HMI tags "xAI"
   "AIx_DB_Level_Use_RTD" : Bool = PLC AIx_DB.Level.Use.RTD AT %DB202.DBX156.0, 1 s
   "AIx_DB_Level_Use_Filter" : Bool = PLC AIx_DB.Level.Use.Filter AT %DB202.DBX156.1, 1 s
   "AIx_DB_Level_Timers_SC_SP" : Int = PLC AIx_DB.Level.Timers.SC.SP AT %DB202.DBW246, 1 s
   "AIx_DB_Level_Timers_NC_SP" : Int = PLC AIx_DB.Level.Timers.NC.SP AT %DB202.DBW240, 1 s
   "AIx_DB_Level_Timers_LL_SP" : Int = PLC AIx_DB.Level.Timers.LL.SP AT %DB202.DBW270, 1 s
   "AIx_DB_Level_Timers_L_SP" : Int = PLC AIx_DB.Level.Timers.L.SP AT %DB202.DBW264, 1 s
   "AIx_DB_Level_Timers_HH_SP" : Int = PLC AIx_DB.Level.Timers.HH.SP AT %DB202.DBW252, 1 s
   "AIx_DB_Level_Timers_H_SP" : Int = PLC AIx_DB.Level.Timers.H.SP AT %DB202.DBW258, 1 s
   "AIx_DB_Level_SP_SC" : Real = PLC AIx_DB.Level.SP.SC AT %DB202.DBD220, 1 s
   "AIx_DB_Level_SP_NC" : Real = PLC AIx_DB.Level.SP.NC AT %DB202.DBD216, 1 s
   "AIx_DB_Level_SP_LL" : Real = PLC AIx_DB.Level.SP.LL AT %DB202.DBD236, 1 s
   "AIx_DB_Level_SP_L" : Real = PLC AIx_DB.Level.SP.L AT %DB202.DBD232, 1 s
   "AIx_DB_Level_SP_HH" : Real = PLC AIx_DB.Level.SP.HH AT %DB202.DBD224, 1 s
   "AIx_DB_Level_SP_H" : Real = PLC AIx_DB.Level.SP.H AT %DB202.DBD228, 1 s
   "AIx_DB_Level_Signal" : Int = PLC AIx_DB.Level.Signal AT %DB202.DBW140, 1 s
   "AIx_DB_Level_RTD_c" : Real = PLC AIx_DB.Level.RTD_c AT %DB202.DBD170, 1 s
   "AIx_DB_Level_Result" : Real = PLC AIx_DB.Level.Result AT %DB202.DBD146, 1 s
   "AIx_DB_Level_Filter_SP" : Real = PLC AIx_DB.Level.Filter.SP AT %DB202.DBD178, 1 s
   "AIx_DB_Level_Converter_Min_Out" : Real = PLC AIx_DB.Level.Converter.Min_Out AT %DB202.DBD208, 1 s
   "AIx_DB_Level_Converter_Min_In" : Real = PLC AIx_DB.Level.Converter.Min_In AT %DB202.DBD200, 1 s
   "AIx_DB_Level_Converter_Max_Out" : Real = PLC AIx_DB.Level.Converter.Max_Out AT %DB202.DBD212, 1 s
   "AIx_DB_Level_Converter_Max_In" : Real = PLC AIx_DB.Level.Converter.Max_In AT %DB202.DBD204, 1 s
   "AIx_DB_Level_CMD_Start_M" : Bool = PLC AIx_DB.Level.CMD.Start_M AT %DB202.DBX150.2, 1 s
   "AIx_DB_Level_CMD_Start_A" : Bool = PLC AIx_DB.Level.CMD.Start_A AT %DB202.DBX150.1, 1 s
   "AIx_DB_Level_CMD_Hand" : Bool = PLC AIx_DB.Level.CMD.Hand AT %DB202.DBX150.0, 1 s
   "AIx_DB_Level_CMD_Alarm" : Bool = PLC AIx_DB.Level.CMD.Alarm AT %DB202.DBX151.0, 1 s
   "AIx_DB_Level_Calibration" : Real = PLC AIx_DB.Level.Calibration AT %DB202.DBD174, 1 s
   "AIx_DB_Level_Alarm" : Word = PLC AIx_DB.Level.Alarm AT %DB202.DBW278, 1 s
   "AIx_DB_FlowMeter_Use_RTD" : Bool = PLC AIx_DB.FlowMeter.Use.RTD AT %DB202.DBX16.0, 1 s
   "AIx_DB_FlowMeter_Use_Filter" : Bool = PLC AIx_DB.FlowMeter.Use.Filter AT %DB202.DBX16.1, 1 s
   "AIx_DB_FlowMeter_Timers_SC_SP" : Int = PLC AIx_DB.FlowMeter.Timers.SC.SP AT %DB202.DBW106, 1 s
   "AIx_DB_FlowMeter_Timers_NC_SP" : Int = PLC AIx_DB.FlowMeter.Timers.NC.SP AT %DB202.DBW100, 1 s
   "AIx_DB_FlowMeter_Timers_LL_SP" : Int = PLC AIx_DB.FlowMeter.Timers.LL.SP AT %DB202.DBW130, 1 s
   "AIx_DB_FlowMeter_Timers_L_SP" : Int = PLC AIx_DB.FlowMeter.Timers.L.SP AT %DB202.DBW124, 1 s
   "AIx_DB_FlowMeter_Timers_HH_SP" : Int = PLC AIx_DB.FlowMeter.Timers.HH.SP AT %DB202.DBW112, 1 s
   "AIx_DB_FlowMeter_Timers_H_SP" : Int = PLC AIx_DB.FlowMeter.Timers.H.SP AT %DB202.DBW118, 1 s
   "AIx_DB_FlowMeter_SP_SC" : Real = PLC AIx_DB.FlowMeter.SP.SC AT %DB202.DBD80, 1 s
   "AIx_DB_FlowMeter_SP_NC" : Real = PLC AIx_DB.FlowMeter.SP.NC AT %DB202.DBD76, 1 s
   "AIx_DB_FlowMeter_SP_LL" : Real = PLC AIx_DB.FlowMeter.SP.LL AT %DB202.DBD96, 1 s
   "AIx_DB_FlowMeter_SP_L" : Real = PLC AIx_DB.FlowMeter.SP.L AT %DB202.DBD92, 1 s
   "AIx_DB_FlowMeter_SP_HH" : Real = PLC AIx_DB.FlowMeter.SP.HH AT %DB202.DBD84, 1 s
   "AIx_DB_FlowMeter_SP_H" : Real = PLC AIx_DB.FlowMeter.SP.H AT %DB202.DBD88, 1 s
   "AIx_DB_FlowMeter_Signal" : Int = PLC AIx_DB.FlowMeter.Signal AT %DB202.DBW0, 1 s
   "AIx_DB_FlowMeter_RTD_c" : Real = PLC AIx_DB.FlowMeter.RTD_c AT %DB202.DBD30, 1 s
   "AIx_DB_FlowMeter_Result" : Real = PLC AIx_DB.FlowMeter.Result AT %DB202.DBD6, 1 s
   "AIx_DB_FlowMeter_Filter_SP" : Real = PLC AIx_DB.FlowMeter.Filter.SP AT %DB202.DBD38, 1 s
   "AIx_DB_FlowMeter_Converter_Min_Out" : Real = PLC AIx_DB.FlowMeter.Converter.Min_Out AT %DB202.DBD68, 1 s
   "AIx_DB_FlowMeter_Converter_Min_In" : Real = PLC AIx_DB.FlowMeter.Converter.Min_In AT %DB202.DBD60, 1 s
   "AIx_DB_FlowMeter_Converter_Max_Out" : Real = PLC AIx_DB.FlowMeter.Converter.Max_Out AT %DB202.DBD72, 1 s
   "AIx_DB_FlowMeter_Converter_Max_In" : Real = PLC AIx_DB.FlowMeter.Converter.Max_In AT %DB202.DBD64, 1 s
   "AIx_DB_FlowMeter_CMD_Start_M" : Bool = PLC AIx_DB.FlowMeter.CMD.Start_M AT %DB202.DBX10.2, 1 s
   "AIx_DB_FlowMeter_CMD_Start_A" : Bool = PLC AIx_DB.FlowMeter.CMD.Start_A AT %DB202.DBX10.1, 1 s
   "AIx_DB_FlowMeter_CMD_Hand" : Bool = PLC AIx_DB.FlowMeter.CMD.Hand AT %DB202.DBX10.0, 1 s
   "AIx_DB_FlowMeter_Calibration" : Real = PLC AIx_DB.FlowMeter.Calibration AT %DB202.DBD34, 1 s
   "AIx_DB_FlowMeter_Alarm" : Word = PLC AIx_DB.FlowMeter.Alarm AT %DB202.DBW138, 1 s

HMI tags "xMotors"
   "Motors_DB_DD_CMD_Start_M" : Bool = PLC Motors_DB.DD.CMD.Start_M AT %DB204.DBX138.2, 1 s
   "Motors_DB_DL_CMD_Hand" : Bool = PLC Motors_DB.DL.CMD.Hand AT %DB204.DBX182.0, 1 s
   "Motors_DB_DL_CMD_Start_M" : Bool = PLC Motors_DB.DL.CMD.Start_M AT %DB204.DBX182.2, 1 s
   "Motors_DB_DL_Res_h" : DInt = PLC Motors_DB.DL.Res_h AT %DB204.DBD212, 1 s
   "Motors_DB_DL_Status" : Int = PLC Motors_DB.DL.Status AT %DB204.DBW186, 1 s
   "Motors_DB_Mix_1_CMD_Force" : Bool = PLC Motors_DB.Mix_1.CMD.Force AT %DB204.DBX6.3, 1 s
   "Motors_DB_Mix_1_CMD_Hand" : Bool = PLC Motors_DB.Mix_1.CMD.Hand AT %DB204.DBX6.0, 1 s
   "Motors_DB_Mix_1_CMD_Service" : Bool = PLC Motors_DB.Mix_1.CMD.Service AT %DB204.DBX6.6, 1 s
   "Motors_DB_Mix_1_CMD_Start_M" : Bool = PLC Motors_DB.Mix_1.CMD.Start_M AT %DB204.DBX6.2, 1 s
   "Motors_DB_Mix_1_FB_KM" : Bool = PLC Motors_DB.Mix_1.FB.KM AT %DB204.DBX14.2, 1 s
   "Motors_DB_Mix_1_FB_QF" : Bool = PLC Motors_DB.Mix_1.FB.QF AT %DB204.DBX14.1, 1 s
   "Motors_DB_Mix_1_FB_Serivce" : Bool = PLC Motors_DB.Mix_1.FB.Serivce AT %DB204.DBX14.3, 1 s
   "Motors_DB_Mix_1_FB_Termo" : Bool = PLC Motors_DB.Mix_1.FB.Termo AT %DB204.DBX14.4, 1 s
   "Motors_DB_Mix_1_Res_h" : DInt = PLC Motors_DB.Mix_1.Res_h AT %DB204.DBD36, 1 s
   "Motors_DB_Mix_1_Status" : Int = PLC Motors_DB.Mix_1.Status AT %DB204.DBW10, 1 s
   "Motors_DB_Mix_1_Use_KM" : Bool = PLC Motors_DB.Mix_1.Use.KM AT %DB204.DBX12.2, 1 s
   "Motors_DB_Mix_1_Use_QF" : Bool = PLC Motors_DB.Mix_1.Use.QF AT %DB204.DBX12.1, 1 s
   "Motors_DB_Mix_1_Use_Serivce" : Bool = PLC Motors_DB.Mix_1.Use.Serivce AT %DB204.DBX12.3, 1 s
   "Motors_DB_Mix_1_Use_Termo" : Bool = PLC Motors_DB.Mix_1.Use.Termo AT %DB204.DBX12.4, 1 s
   "Motors_DB_Mix_1_Wait_Off_Now" : Int = PLC Motors_DB.Mix_1.Wait_Off.Now AT %DB204.DBW26, 1 s
   "Motors_DB_Mix_1_Wait_Off_SP" : Int = PLC Motors_DB.Mix_1.Wait_Off.SP AT %DB204.DBW24, 1 s
   "Motors_DB_Mix_1_Wait_On_Now" : Int = PLC Motors_DB.Mix_1.Wait_On.Now AT %DB204.DBW20, 1 s
   "Motors_DB_Mix_1_Wait_On_SP" : Int = PLC Motors_DB.Mix_1.Wait_On.SP AT %DB204.DBW18, 1 s
   "Motors_DB_Mix_2_CMD_Hand" : Bool = PLC Motors_DB.Mix_2.CMD.Hand AT %DB204.DBX50.0, 1 s
   "Motors_DB_Mix_2_CMD_Start_M" : Bool = PLC Motors_DB.Mix_2.CMD.Start_M AT %DB204.DBX50.2, 1 s
   "Motors_DB_Mix_2_Res_h" : DInt = PLC Motors_DB.Mix_2.Res_h AT %DB204.DBD80, 1 s
   "Motors_DB_Mix_2_Status" : Int = PLC Motors_DB.Mix_2.Status AT %DB204.DBW54, 1 s
   "Motors_DB_Mix_3_CMD_Hand" : Bool = PLC Motors_DB.Mix_3.CMD.Hand AT %DB204.DBX94.0, 1 s
   "Motors_DB_Mix_3_CMD_Start_M" : Bool = PLC Motors_DB.Mix_3.CMD.Start_M AT %DB204.DBX94.2, 1 s
   "Motors_DB_Mix_3_Res_h" : DInt = PLC Motors_DB.Mix_3.Res_h AT %DB204.DBD124, 1 s
   "Motors_DB_Mix_3_Status" : Int = PLC Motors_DB.Mix_3.Status AT %DB204.DBW98, 1 s
   "Motors_DB_Mix_2_CMD_Force" : Bool = PLC Motors_DB.Mix_2.CMD.Force AT %DB204.DBX50.3, 1 s
   "Motors_DB_Mix_2_CMD_Service" : Bool = PLC Motors_DB.Mix_2.CMD.Service AT %DB204.DBX50.6, 1 s
   "Motors_DB_Mix_2_Use_QF" : Bool = PLC Motors_DB.Mix_2.Use.QF AT %DB204.DBX56.1, 1 s
   "Motors_DB_Mix_2_Use_KM" : Bool = PLC Motors_DB.Mix_2.Use.KM AT %DB204.DBX56.2, 1 s
   "Motors_DB_Mix_2_Use_Serivce" : Bool = PLC Motors_DB.Mix_2.Use.Serivce AT %DB204.DBX56.3, 1 s
   "Motors_DB_Mix_2_Use_Termo" : Bool = PLC Motors_DB.Mix_2.Use.Termo AT %DB204.DBX56.4, 1 s
   "Motors_DB_Mix_2_FB_QF" : Bool = PLC Motors_DB.Mix_2.FB.QF AT %DB204.DBX58.1, 1 s
   "Motors_DB_Mix_2_FB_KM" : Bool = PLC Motors_DB.Mix_2.FB.KM AT %DB204.DBX58.2, 1 s
   "Motors_DB_Mix_2_FB_Serivce" : Bool = PLC Motors_DB.Mix_2.FB.Serivce AT %DB204.DBX58.3, 1 s
   "Motors_DB_Mix_2_FB_Termo" : Bool = PLC Motors_DB.Mix_2.FB.Termo AT %DB204.DBX58.4, 1 s
   "Motors_DB_Mix_2_Alarm" : Word = PLC Motors_DB.Mix_2.Alarm AT %DB204.DBW78, 1 s
   "Motors_DB_Mix_2_Wait_On_SP" : Int = PLC Motors_DB.Mix_2.Wait_On.SP AT %DB204.DBW62, 1 s
   "Motors_DB_Mix_2_Wait_On_Now" : Int = PLC Motors_DB.Mix_2.Wait_On.Now AT %DB204.DBW64, 1 s
   "Motors_DB_Mix_2_Wait_Off_SP" : Int = PLC Motors_DB.Mix_2.Wait_Off.SP AT %DB204.DBW68, 1 s
   "Motors_DB_Mix_2_Wait_Off_Now" : Int = PLC Motors_DB.Mix_2.Wait_Off.Now AT %DB204.DBW70, 1 s
   "Motors_DB_Mix_1_Alarm" : Word = PLC Motors_DB.Mix_1.Alarm AT %DB204.DBW34, 1 s
   "Motors_DB_Mix_3_CMD_Start_A" : Bool = PLC Motors_DB.Mix_3.CMD.Start_A AT %DB204.DBX94.1, 1 s
   "Motors_DB_Mix_3_CMD_Force" : Bool = PLC Motors_DB.Mix_3.CMD.Force AT %DB204.DBX94.3, 1 s
   "Motors_DB_Mix_3_CMD_Service" : Bool = PLC Motors_DB.Mix_3.CMD.Service AT %DB204.DBX94.6, 1 s
   "Motors_DB_Mix_3_Use_QF" : Bool = PLC Motors_DB.Mix_3.Use.QF AT %DB204.DBX100.1, 1 s
   "Motors_DB_Mix_3_Use_KM" : Bool = PLC Motors_DB.Mix_3.Use.KM AT %DB204.DBX100.2, 1 s
   "Motors_DB_Mix_3_Use_Serivce" : Bool = PLC Motors_DB.Mix_3.Use.Serivce AT %DB204.DBX100.3, 1 s
   "Motors_DB_Mix_3_Use_Termo" : Bool = PLC Motors_DB.Mix_3.Use.Termo AT %DB204.DBX100.4, 1 s
   "Motors_DB_Mix_3_FB_QF" : Bool = PLC Motors_DB.Mix_3.FB.QF AT %DB204.DBX102.1, 1 s
   "Motors_DB_Mix_3_FB_KM" : Bool = PLC Motors_DB.Mix_3.FB.KM AT %DB204.DBX102.2, 1 s
   "Motors_DB_Mix_3_FB_Serivce" : Bool = PLC Motors_DB.Mix_3.FB.Serivce AT %DB204.DBX102.3, 1 s
   "Motors_DB_Mix_3_FB_Termo" : Bool = PLC Motors_DB.Mix_3.FB.Termo AT %DB204.DBX102.4, 1 s
   "Motors_DB_Mix_3_Alarm" : Word = PLC Motors_DB.Mix_3.Alarm AT %DB204.DBW122, 1 s
   "Motors_DB_Mix_3_Wait_On_SP" : Int = PLC Motors_DB.Mix_3.Wait_On.SP AT %DB204.DBW106, 1 s
   "Motors_DB_Mix_3_Wait_On_Now" : Int = PLC Motors_DB.Mix_3.Wait_On.Now AT %DB204.DBW108, 1 s
   "Motors_DB_Mix_3_Wait_Off_SP" : Int = PLC Motors_DB.Mix_3.Wait_Off.SP AT %DB204.DBW112, 1 s
   "Motors_DB_Mix_3_Wait_Off_Now" : Int = PLC Motors_DB.Mix_3.Wait_Off.Now AT %DB204.DBW114, 1 s
   "Motors_DB_DD_CMD_Hand" : Bool = PLC Motors_DB.DD.CMD.Hand AT %DB204.DBX138.0, 1 s
   "Motors_DB_DD_CMD_Force" : Bool = PLC Motors_DB.DD.CMD.Force AT %DB204.DBX138.3, 1 s
   "Motors_DB_DD_CMD_Service" : Bool = PLC Motors_DB.DD.CMD.Service AT %DB204.DBX138.6, 1 s
   "Motors_DB_DD_Use_QF" : Bool = PLC Motors_DB.DD.Use.QF AT %DB204.DBX144.1, 1 s
   "Motors_DB_DD_Use_KM" : Bool = PLC Motors_DB.DD.Use.KM AT %DB204.DBX144.2, 1 s
   "Motors_DB_DD_Use_Serivce" : Bool = PLC Motors_DB.DD.Use.Serivce AT %DB204.DBX144.3, 1 s
   "Motors_DB_DD_Use_Termo" : Bool = PLC Motors_DB.DD.Use.Termo AT %DB204.DBX144.4, 1 s
   "Motors_DB_DD_FB_QF" : Bool = PLC Motors_DB.DD.FB.QF AT %DB204.DBX146.1, 1 s
   "Motors_DB_DD_FB_KM" : Bool = PLC Motors_DB.DD.FB.KM AT %DB204.DBX146.2, 1 s
   "Motors_DB_DD_FB_Serivce" : Bool = PLC Motors_DB.DD.FB.Serivce AT %DB204.DBX146.3, 1 s
   "Motors_DB_DD_FB_Termo" : Bool = PLC Motors_DB.DD.FB.Termo AT %DB204.DBX146.4, 1 s
   "Motors_DB_DD_Alarm" : Word = PLC Motors_DB.DD.Alarm AT %DB204.DBW166, 1 s
   "Motors_DB_DD_Wait_On_SP" : Int = PLC Motors_DB.DD.Wait_On.SP AT %DB204.DBW150, 1 s
   "Motors_DB_DD_Wait_On_Now" : Int = PLC Motors_DB.DD.Wait_On.Now AT %DB204.DBW152, 1 s
   "Motors_DB_DD_Wait_Off_SP" : Int = PLC Motors_DB.DD.Wait_Off.SP AT %DB204.DBW156, 1 s
   "Motors_DB_DD_Wait_Off_Now" : Int = PLC Motors_DB.DD.Wait_Off.Now AT %DB204.DBW158, 1 s
   "Motors_DB_DL_CMD_Force" : Bool = PLC Motors_DB.DL.CMD.Force AT %DB204.DBX182.3, 1 s
   "Motors_DB_DL_CMD_Service" : Bool = PLC Motors_DB.DL.CMD.Service AT %DB204.DBX182.6, 1 s
   "Motors_DB_DL_Use_QF" : Bool = PLC Motors_DB.DL.Use.QF AT %DB204.DBX188.1, 1 s
   "Motors_DB_DL_Use_KM" : Bool = PLC Motors_DB.DL.Use.KM AT %DB204.DBX188.2, 1 s
   "Motors_DB_DL_Use_Serivce" : Bool = PLC Motors_DB.DL.Use.Serivce AT %DB204.DBX188.3, 1 s
   "Motors_DB_DL_Use_Termo" : Bool = PLC Motors_DB.DL.Use.Termo AT %DB204.DBX188.4, 1 s
   "Motors_DB_DL_FB_QF" : Bool = PLC Motors_DB.DL.FB.QF AT %DB204.DBX190.1, 1 s
   "Motors_DB_DL_FB_KM" : Bool = PLC Motors_DB.DL.FB.KM AT %DB204.DBX190.2, 1 s
   "Motors_DB_DL_FB_Serivce" : Bool = PLC Motors_DB.DL.FB.Serivce AT %DB204.DBX190.3, 1 s
   "Motors_DB_DL_FB_Termo" : Bool = PLC Motors_DB.DL.FB.Termo AT %DB204.DBX190.4, 1 s
   "Motors_DB_DL_Alarm" : Word = PLC Motors_DB.DL.Alarm AT %DB204.DBW210, 1 s
   "Motors_DB_DL_Wait_On_SP" : Int = PLC Motors_DB.DL.Wait_On.SP AT %DB204.DBW194, 1 s
   "Motors_DB_DL_Wait_On_Now" : Int = PLC Motors_DB.DL.Wait_On.Now AT %DB204.DBW196, 1 s
   "Motors_DB_DL_Wait_Off_SP" : Int = PLC Motors_DB.DL.Wait_Off.SP AT %DB204.DBW200, 1 s
   "Motors_DB_DL_Wait_Off_Now" : Int = PLC Motors_DB.DL.Wait_Off.Now AT %DB204.DBW202, 1 s
   "Motors_DB_Vibro_CMD_Force" : Bool = PLC Motors_DB.Vibro.CMD.Force AT %DB204.DBX226.3, 1 s
   "Motors_DB_Vibro_CMD_Service" : Bool = PLC Motors_DB.Vibro.CMD.Service AT %DB204.DBX226.6, 1 s
   "Motors_DB_Vibro_Use_QF" : Bool = PLC Motors_DB.Vibro.Use.QF AT %DB204.DBX232.1, 1 s
   "Motors_DB_Vibro_Use_KM" : Bool = PLC Motors_DB.Vibro.Use.KM AT %DB204.DBX232.2, 1 s
   "Motors_DB_Vibro_Use_Serivce" : Bool = PLC Motors_DB.Vibro.Use.Serivce AT %DB204.DBX232.3, 1 s
   "Motors_DB_Vibro_Use_Termo" : Bool = PLC Motors_DB.Vibro.Use.Termo AT %DB204.DBX232.4, 1 s
   "Motors_DB_Vibro_FB_QF" : Bool = PLC Motors_DB.Vibro.FB.QF AT %DB204.DBX234.1, 1 s
   "Motors_DB_Vibro_FB_KM" : Bool = PLC Motors_DB.Vibro.FB.KM AT %DB204.DBX234.2, 1 s
   "Motors_DB_Vibro_FB_Serivce" : Bool = PLC Motors_DB.Vibro.FB.Serivce AT %DB204.DBX234.3, 1 s
   "Motors_DB_Vibro_FB_Termo" : Bool = PLC Motors_DB.Vibro.FB.Termo AT %DB204.DBX234.4, 1 s
   "Motors_DB_Vibro_CMD_Start_M" : Bool = PLC Motors_DB.Vibro.CMD.Start_M AT %DB204.DBX226.2, 1 s
   "Motors_DB_Vibro_CMD_Hand" : Bool = PLC Motors_DB.Vibro.CMD.Hand AT %DB204.DBX226.0, 1 s
   "Motors_DB_Vibro_Alarm" : Word = PLC Motors_DB.Vibro.Alarm AT %DB204.DBW254, 1 s
   "Motors_DB_Vibro_Wait_On_SP" : Int = PLC Motors_DB.Vibro.Wait_On.SP AT %DB204.DBW238, 1 s
   "Motors_DB_Vibro_Wait_On_Now" : Int = PLC Motors_DB.Vibro.Wait_On.Now AT %DB204.DBW240, 1 s
   "Motors_DB_Vibro_Wait_Off_SP" : Int = PLC Motors_DB.Vibro.Wait_Off.SP AT %DB204.DBW244, 1 s
   "Motors_DB_Vibro_Wait_Off_Now" : Int = PLC Motors_DB.Vibro.Wait_Off.Now AT %DB204.DBW246, 1 s

HMI tags "xValve"
   "Micro_DB_KC1_Status" : Int = PLC Micro_DB.KC1.Status AT %DB207.DBW8, 1 s
   "Micro_DB_KC1_Start_M" : Bool = PLC Micro_DB.KC1.Start_M AT %DB207.DBX6.1, 1 s
   "Micro_DB_KC1_Hand" : Bool = PLC Micro_DB.KC1.Hand AT %DB207.DBX6.0, 1 s
   "Micro_DB_KC1_CMD" : Bool = PLC Micro_DB.KC1.CMD AT %DB207.DBX2.0, 1 s
   "Micro_DB_KC1_Alarm" : Bool = PLC Micro_DB.KC1.Alarm AT %DB207.DBX4.0, 1 s
   "Micro_DB_KC1_No_FB" : Bool = PLC Micro_DB.KC1.No_FB AT %DB207.DBX6.2, 1 s
   "Micro_DB_KC1_Wait_Off_SP" : Int = PLC Micro_DB.KC1.Wait_Off.SP AT %DB207.DBW16, 1 s
   "Micro_DB_KC1_Wait_On_SP" : Int = PLC Micro_DB.KC1.Wait_On.SP AT %DB207.DBW10, 1 s

discrete alarms
   1: 'Авария - Сработал датчик протока', class Errors, trigger "Logick_DB_Alarm" bit 0
   2: 'Авария - Низкий уровень в бункере', class Errors, trigger "Logick_DB_Alarm" bit 1
   3: 'Внешний остнова / Перелив', class Errors, trigger "Logick_DB_Alarm" bit 2
   4: 'Предупреждение - Нет готовности пнемотранспортёра', class Errors, trigger "Logick_DB_Alarm" bit 3
   5: 'Уровень - Обрыв датчика', class Errors, trigger "AIx_DB_Level_Alarm" bit 0
   6: 'Уровень - Короткое замыкание', class Errors, trigger "AIx_DB_Level_Alarm" bit 1
   7: 'Уровень - Аварийно высокий уровнь', class Errors, trigger "AIx_DB_Level_Alarm" bit 2
   8: 'Уровень - Высокий уровень', class Errors, trigger "AIx_DB_Level_Alarm" bit 3
   9: 'Уровень - Низкий уровень', class Errors, trigger "AIx_DB_Level_Alarm" bit 4
   10: 'Уровень - Аварийно низкий уровень', class Errors, trigger "AIx_DB_Level_Alarm" bit 5
   11: 'Расходомер - Обрыв датчика', class Errors, trigger "AIx_DB_FlowMeter_Alarm" bit 0
   12: 'Расходомер - Короткое замыкание', class Errors, trigger "AIx_DB_FlowMeter_Alarm" bit 1
   13: 'Расходомер - Аварийно высокий поток', class Errors, trigger "AIx_DB_FlowMeter_Alarm" bit 2
   14: 'Расходомер - Высокий поток', class Errors, trigger "AIx_DB_FlowMeter_Alarm" bit 3
   15: 'Расходомер - Низкий поток', class Errors, trigger "AIx_DB_FlowMeter_Alarm" bit 4
   16: 'Расходомер - Аварийно низкий поток', class Errors, trigger "AIx_DB_FlowMeter_Alarm" bit 5
   17: 'Мешалка 1 - Выбило защитный автомат', class Errors, trigger "Motors_DB_Mix_1_Alarm" bit 0
   18: 'Мешалка 1 - Ошибка при запуске', class Errors, trigger "Motors_DB_Mix_1_Alarm" bit 1
   19: 'Мешалка 1 - Ошибка при останове', class Errors, trigger "Motors_DB_Mix_1_Alarm" bit 2
   20: 'Мешалка 1 - Сработало реле безопасности', class Errors, trigger "Motors_DB_Mix_1_Alarm" bit 3
   21: 'Мешалка 1 - Общая блокировка', class Errors, trigger "Motors_DB_Mix_1_Alarm" bit 4
   22: 'Мешалка 1 - Перегрев двигателя', class Errors, trigger "Motors_DB_Mix_1_Alarm" bit 5
   23: 'Мешалка 2 - Выбило защитный автомат', class Errors, trigger "Motors_DB_Mix_2_Alarm" bit 0
   24: 'Мешалка 2 - Ошибка при запуске', class Errors, trigger "Motors_DB_Mix_2_Alarm" bit 1
   25: 'Мешалка 2 - Ошибка при останове', class Errors, trigger "Motors_DB_Mix_2_Alarm" bit 2
   26: 'Мешалка 2 - Сработало реле безопасности', class Errors, trigger "Motors_DB_Mix_2_Alarm" bit 3
   27: 'Мешалка 2 - Общая блокировка', class Errors, trigger "Motors_DB_Mix_2_Alarm" bit 4
   28: 'Мешалка 2 - Перегрев двигателя', class Errors, trigger "Motors_DB_Mix_2_Alarm" bit 5
   29: 'Мешалка 3 - Выбило защитный автомат', class Errors, trigger "Motors_DB_Mix_3_Alarm" bit 0
   30: 'Мешалка 3 - Ошибка при запуске', class Errors, trigger "Motors_DB_Mix_3_Alarm" bit 1
   31: 'Мешалка 3 - Ошибка при останове', class Errors, trigger "Motors_DB_Mix_3_Alarm" bit 2
   32: 'Мешалка 3 - Сработало реле безопасности', class Errors, trigger "Motors_DB_Mix_3_Alarm" bit 3
   33: 'Мешалка 3 - Общая блокировка', class Errors, trigger "Motors_DB_Mix_3_Alarm" bit 4
   34: 'Мешалка 3 - Перегрев двигателя', class Errors, trigger "Motors_DB_Mix_3_Alarm" bit 5
   35: 'Сухой дозатор - Выбило защитный автомат', class Errors, trigger "Motors_DB_DD_Alarm" bit 0
   36: 'Сухой дозатор - Ошибка при запуске', class Errors, trigger "Motors_DB_DD_Alarm" bit 1
   37: 'Сухой дозатор - Ошибка при останове', class Errors, trigger "Motors_DB_DD_Alarm" bit 2
   38: 'Сухой дозатор - Сработало реле безопасности', class Errors, trigger "Motors_DB_DD_Alarm" bit 3
   39: 'Сухой дозатор - Общая блокировка', class Errors, trigger "Motors_DB_DD_Alarm" bit 4
   40: 'Сухой дозатор - Перегрев двигателя', class Errors, trigger "Motors_DB_DD_Alarm" bit 5
   41: 'Жидкий дозатор - Устройство не готово', class Errors, trigger "Motors_DB_DL_Alarm" bit 0
   42: 'Жидкий дозатор - Ошибка при запуске', class Errors, trigger "Motors_DB_DL_Alarm" bit 1
   43: 'Жидкий дозатор - Ошибка при останове', class Errors, trigger "Motors_DB_DL_Alarm" bit 2
   44: 'Жидкий дозатор - Сработало реле безопасности', class Errors, trigger "Motors_DB_DL_Alarm" bit 3
   45: 'Жидкий дозатор - Общая блокировка', class Errors, trigger "Motors_DB_DL_Alarm" bit 4
   46: 'Жидкий дозатор - Перегрев двигателя', class Errors, trigger "Motors_DB_DL_Alarm" bit 5
   47: 'Вибратор - Устройство не готово', class Errors, trigger "Motors_DB_Vibro_Alarm" bit 0
   48: 'Вибратор - Ошибка при запуске', class Errors, trigger "Motors_DB_Vibro_Alarm" bit 1
   49: 'Вибратор - Ошибка при останове', class Errors, trigger "Motors_DB_Vibro_Alarm" bit 2
   50: 'Вибратор - Сработало реле безопасности', class Errors, trigger "Motors_DB_Vibro_Alarm" bit 3
   51: 'Вибратор - Общая блокировка', class Errors, trigger "Motors_DB_Vibro_Alarm" bit 4
   52: 'Вибратор - Перегрев двигателя', class Errors, trigger "Motors_DB_Vibro_Alarm" bit 5

text list "Hand": 0 'Авто'; 1 'Ручной'

text list "настройки": 0 'Настройки >>'; 1 'Настройки <<'

graphic list "Motor": 0 'm_off_1'; 1 'm_on_1'; 2..8 'm_wait_1'; 9..1000 'm_alarm_1'

graphic list "Pump": 0 'p_off'; 1 'p_on'; 2..8 'p_wait'; 9..1000 'p_alarm'

graphic list "Valve": 0 'v_off'; 1 'v_on'; 2..8 'v_wait'; 9..1000 'v_alarm'

graphic list "L_1": 0 'L_1_off'; 1 'L_1_on'; 2..8 'L_1_wait'; 9..1000 'L_1_alarm'

graphic list "L_2": 0 'L_2_off'; 1 'L_2_on'; 2..8 'L_2_wait'; 9..1000 'L_2_alarm'

graphic list "Led": 0 'no_alarm_led'; 1 'alarm_led'

graphic list "Alarm": 0 'no_alarm_1'; 1 'alarm'

graphic list "ON_OFF": 0 'off_toggle'; 1 'on_toggle'

graphic list "ok": 0 'check_box_off'; 1 'check_box_on'

graphic list "Status": 0 'sys_x'; 1 'sys_check-mark'; 2 'z2use'; 3..99 'alarm_on'

graphic list "Vibro": 0 'b_1'; 1 'b_4'; 2..4 'b_2'; 5..1000 'b_3'

screen "Root screen" 800x480, template "Main"
   GraphicView "Graphic view_3" at 5,58 size 40x183; Picture "Graphic_5"
   GraphicView "Graphic view_4" at 324,272 size 164x200; Picture "h2o_1"
   GraphicView "Graphic view_2" at 166,272 size 164x200; Picture "h2o_1"
   Rectangle "Rectangle_8" at 543,104 size 175x115
      Visibility <- "Any_Hand"
      Appearance <- "Any_Hand"
   GraphicView "Graphic view_7" at 5,21 size 40x40; Picture "Graphic_6"
   GraphicView "Graphic view_5" at 41,21 size 200x40; Picture "Graphic_4"
   GraphicView "Graphic view_6" at 33,93 size 214x40; Picture "Graphic_4"
   Bar "Bar_1" at 440,235 size 85x240; Unit %; MinimumValue 0; MaximumValue 100
      ProcessValue <- "AIx_DB_Level_Result"
   GraphicView "Graphic view_1" at 8,272 size 164x200; Picture "h2o_1"
   GraphicIOField "Graphic I/O field_2" at 240,157 size 50x93; PictureList "Motor"
      ProcessValue <- "Motors_DB_Mix_2_Status"
   GraphicIOField "Graphic I/O field_3" at 415,157 size 50x93; PictureList "Motor"
      ProcessValue <- "Motors_DB_Mix_3_Status"
   GraphicIOField "Graphic I/O field_4" at 237,86 size 50x50; PictureList "Pump"
      ProcessValue <- "Motors_DB_DL_Status"
   Rectangle "Rectangle_4" at 5,62 size 40x100
      Visibility <- "CONFIG_Config_Use_DL"
   Line "Line_1" at 4,63 size 40x40
      Visibility <- "CONFIG_Config_Use_DL"
   Line "Line_2" at 4,92 size 40x40
      Visibility <- "CONFIG_Config_Use_DL"
   Line "Line_3" at 4,122 size 40x40
      Visibility <- "CONFIG_Config_Use_DL"
   Line "Line_4" at 5,62 size 40x40
      Visibility <- "CONFIG_Config_Use_DL"
   Line "Line_5" at 5,92 size 40x40
      Visibility <- "CONFIG_Config_Use_DL"
   Line "Line_6" at 5,122 size 40x40
      Visibility <- "CONFIG_Config_Use_DL"
   GraphicIOField "Graphic I/O field_5" at 237,2 size 50x50; PictureList "Valve"
      ProcessValue <- "Micro_DB_KC1_Status"
   IOField "I/O field_1" at 88,24 size 103x32; FormatPattern 9999.9
      ProcessValue <- "AIx_DB_FlowMeter_Result"
   TextField "Text field_1" at 154,27 size 34x23; Text 'л/ч'
   TextField "Text field_2" at 85,2 size 107x23; Text 'Расходомер'
   TextField "Text field_3" at 241,50 size 37x23; Text 'КС1'
   GraphicIOField "Graphic I/O field_1" at 65,157 size 50x93; PictureList "Motor"
      ProcessValue <- "Motors_DB_Mix_1_Status"
   GraphicIOField "Graphic I/O field_7" at 190,425 size 150x40; PictureList "L_1"
      Visibility <- "Mix_2_Clock"
      ProcessValue <- "Motors_DB_Mix_2_Status"
   GraphicIOField "Graphic I/O field_8" at 365,425 size 150x40; PictureList "L_1"
      Visibility <- "Mix_3_Clock"
      ProcessValue <- "Motors_DB_Mix_3_Status"
   GraphicIOField "Graphic I/O field_10" at 190,425 size 150x40; PictureList "L_2"
      Visibility <- "Mix_2_Clock"
      ProcessValue <- "Motors_DB_Mix_2_Status"
   GraphicIOField "Graphic I/O field_11" at 365,425 size 150x40; PictureList "L_2"
      Visibility <- "Mix_3_Clock"
      ProcessValue <- "Motors_DB_Mix_3_Status"
   GraphicIOField "Graphic I/O field_6" at 15,425 size 150x40; PictureList "L_1"
      Visibility <- "Mix_1_Clock"
      ProcessValue <- "Motors_DB_Mix_1_Status"
   GraphicIOField "Graphic I/O field_9" at 15,425 size 150x40; PictureList "L_2"
      Visibility <- "Mix_1_Clock"
      ProcessValue <- "Motors_DB_Mix_1_Status"
   GraphicIOField "Graphic I/O field_12" at 495,168 size 30x40; PictureList "Led"
      ProcessValue <- "AIx_DB_Level_CMD_Alarm"
   TextField "Text field_4" at 439,6 size 218x27; Text 'система дозирования'
   TextField "Text field_5" at 434,27 size 227x72; Text 'PolyMix'
   Button "Button_8" at 543,238 size 175x60; TextOff 'Авто'
      on Click: SetBit("Logick_DB_Start")
      Appearance <- "Logick_DB_Start"
   Button "Button_9" at 543,326 size 175x60; TextOff 'Стоп'
      on Click: ResetBit("Logick_DB_Start")
   Button "Button_10" at 543,415 size 175x60; TextOff 'Ручной'; Authorization "Operator"
      on Click: InvertBit("Logick_DB_Hand")
      Appearance <- "Logick_DB_Hand"
   Button "Button_11" at 236,2 size 51x52; TextOff 'Text'; Authorization "Operator"
      on Click: InvertBit("Micro_DB_KC1_Start_M")
      Visibility <- "Micro_DB_KC1_Hand"
   Button "Button_12" at 236,86 size 51x52; TextOff 'Text'; Authorization "Operator"
      on Click: InvertBit("Motors_DB_DL_CMD_Start_M")
      Visibility <- "Motors_DB_DL_CMD_Hand"
   Button "Button_13" at 64,155 size 51x79; TextOff 'Text'; Authorization "Operator"
      on Click: InvertBit("Motors_DB_Mix_1_CMD_Start_M")
      Visibility <- "Motors_DB_Mix_1_CMD_Hand"
   Button "Button_14" at 15,422 size 153x43; TextOff 'Text'; Authorization "Operator"
      on Click: InvertBit("Motors_DB_Mix_1_CMD_Start_M")
      Visibility <- "Motors_DB_Mix_1_CMD_Hand"
   Button "Button_15" at 241,155 size 51x79; TextOff 'Text'; Authorization "Operator"
      on Click: InvertBit("Motors_DB_Mix_2_CMD_Start_M")
      Visibility <- "Motors_DB_Mix_2_CMD_Hand"
   Button "Button_16" at 192,422 size 153x43; TextOff 'Text'; Authorization "Operator"
      on Click: InvertBit("Motors_DB_Mix_2_CMD_Start_M")
      Visibility <- "Motors_DB_Mix_2_CMD_Hand"
   Button "Button_17" at 416,155 size 51x79; TextOff 'Text'; Authorization "Operator"
      on Click: InvertBit("Motors_DB_Mix_3_CMD_Start_M")
      Visibility <- "Motors_DB_Mix_3_CMD_Hand"
   Button "Button_18" at 367,422 size 153x43; TextOff 'Text'; Authorization "Operator"
      on Click: InvertBit("Motors_DB_Mix_3_CMD_Start_M")
      Visibility <- "Motors_DB_Mix_3_CMD_Hand"
   IOField "I/O field_2" at 288,85 size 96x32; FormatPattern 9999999
      Visibility <- "Logick_DB_Hand"
      ProcessValue <- "Motors_DB_DL_Res_h"
   TextField "Text field_6" at 363,89 size 15x23; Text 'ч'
      Visibility <- "Logick_DB_Hand"
   IOField "I/O field_3" at 115,155 size 96x32; FormatPattern 9999999
      ProcessValue <- "Motors_DB_Mix_1_Res_h"
      Visibility <- "Logick_DB_Hand"
   TextField "Text field_7" at 190,158 size 15x23; Text 'ч'
      Visibility <- "Logick_DB_Hand"
   IOField "I/O field_4" at 289,155 size 96x32; FormatPattern 9999999
      ProcessValue <- "Motors_DB_Mix_2_Res_h"
      Visibility <- "Logick_DB_Hand"
   TextField "Text field_8" at 364,158 size 15x23; Text 'ч'
      Visibility <- "Logick_DB_Hand"
   IOField "I/O field_5" at 416,123 size 96x32; FormatPattern 9999999
      ProcessValue <- "Motors_DB_Mix_3_Res_h"
      Visibility <- "Logick_DB_Hand"
   TextField "Text field_9" at 491,126 size 15x23; Text 'ч'
      Visibility <- "Logick_DB_Hand"
   TextField "Text field_10" at 547,111 size 169x99; Text 'Внимание! Часть устройств в ручном режиме. Корректная работа невозможна.'
      Visibility <- "Any_Hand"
      Appearance <- "Any_Hand"
   Rectangle "Rectangle_9" at 121,103 size 34x18
      Appearance <- "DIx_DB_Dry_Run_Signal"
   IOField "I/O field_8" at 467,208 size 58x27; Authorization "Operator"; FormatPattern 999
      ProcessValue <- "AIx_DB_Level_Result"
      Appearance <- "AIx_DB_Level_CMD_Alarm"
   TextField "Text field_11" at 501,210 size 24x23; Text '%'
   IOField "I/O field_6" at 61,52 size 160x32; FormatPattern 99999999999999
      ProcessValue <- "FlowMeter_DB_Full"
      Visibility <- "Logick_DB_Hand"
   TextField "Text field_12" at 205,56 size 15x23; Text 'л'
      Visibility <- "Logick_DB_Hand"
   Rectangle "Rectangle_2" at 27,84 size 358x58
      Visibility <- "CONFIG_Config_Use_DD"
   GraphicView "Graphic view_8" at 28,128 size 40x108; Picture "Graphic_5"
      Visibility <- "CONFIG_Config_Use_DD"
   Rectangle "Rectangle_3" at 37,112 size 255x25
      Visibility <- "CONFIG_Config_Use_DD"
      Appearance <- "Motors_DB_DD_Status"
   Line "Line_9" at 38,113 size 38x23
      Visibility <- "CONFIG_Config_Use_DD"
   Line "Line_10" at 73,113 size 38x23
      Visibility <- "CONFIG_Config_Use_DD"
   Line "Line_11" at 110,113 size 38x23
      Visibility <- "CONFIG_Config_Use_DD"
   Line "Line_12" at 145,113 size 38x23
      Visibility <- "CONFIG_Config_Use_DD"
   Line "Line_13" at 182,113 size 38x23
      Visibility <- "CONFIG_Config_Use_DD"
   Line "Line_14" at 217,113 size 38x23
      Visibility <- "CONFIG_Config_Use_DD"
   Line "Line_15" at 256,113 size 38x23
      Visibility <- "CONFIG_Config_Use_DD"
   GraphicIOField "Graphic I/O field_13" at 290,38 size 100x100; PictureList "Vibro"
      ProcessValue <- "Motors_DB_Vibro_Status"
      Visibility <- "CONFIG_Config_Use_DD"
   Rectangle "Rectangle_10" at 292,113 size 96x23
      Visibility <- "CONFIG_Config_Use_DD"
      Appearance <- "DIx_DB_DD_LLS_Signal"
   Button "Button_1" at 289,38 size 98x74; TextOff 'Text'
      on Click: InvertBit("Motors_DB_Vibro_CMD_Start_M")
      Visibility <- "CONFIG_Config_Use_DD"
   Button "Button_2" at 38,111 size 256x26; TextOff 'Text'
      on Click: InvertBit("Motors_DB_DD_CMD_Start_M")
      Visibility <- "CONFIG_Config_Use_DD"
   Rectangle "Rectangle_11" at 22,260 size 406x145
      Visibility <- "Any_DB_Level_View"
   TextField "Text field_13" at 107,269 size 235x29; Text 'Низкий уровень в баке'
      Visibility <- "AIx_DB_Level_Alarms_LL"
   TextField "Text field_14" at 107,301 size 175x27; Text 'остановка через:'
      Visibility <- "Any_DB_Level_View"
   IOField "I/O field_7" at 286,301 size 37x32; FormatPattern 99
      Visibility <- "Any_DB_Level_View"
      ProcessValue <- "Any_DB_Level_M"
   TextField "Text field_15" at 324,302 size 19x27; Text 'м'
      Visibility <- "Any_DB_Level_View"
   Button "Button_3" at 151,350 size 150x32; TextOff 'Игнорировать'
      on Click: SetBit("Logick_DB_Level_CMD")
      Visibility <- "Any_DB_Level_View"
      Appearance <- "Logick_DB_Level_CMD"
   TextField "Text field_16" at 99,269 size 249x29; Text 'Высокий уровень в баке'
      Visibility <- "AIx_DB_Level_Alarms_HH"
   Group "Group" at 22,260 size 406x145
   Button "Button_5" at 151,351 size 150x32; TextOff 'Игнорировать'
      on Click: SetBit("Logick_DB_DD_CMD")
      Appearance <- "Logick_DB_DD_CMD"
      Visibility <- "Any_DB_DD_View"
   Button "Button_4" at 151,350 size 150x32; TextOff 'Игнорировать'
      on Click: SetBit("Logick_DB_DD_CMD")
      Appearance <- "Logick_DB_DD_CMD"
      Visibility <- "Any_DB_DD_View"
   Rectangle "Rectangle_12" at 22,260 size 406x145
      Visibility <- "Any_DB_DD_View"
   TextField "Text field_18" at 324,302 size 19x27; Text 'м'
      Visibility <- "Any_DB_DD_View"
   IOField "I/O field_9" at 286,301 size 37x32; FormatPattern 99
      Visibility <- "Any_DB_DD_View"
      ProcessValue <- "Any_DB_Flow_M"
   TextField "Text field_17" at 107,301 size 175x27; Text 'остановка через:'
      Visibility <- "Any_DB_DD_View"
   TextField "Text field_19" at 77,271 size 309x27; Text 'Нет протока / Низкий уровень'
      Visibility <- "Any_DB_DD_View"

screen "Alarms" 800x480, template "Main"
   AlarmView "Alarm view_1" at 4,3 size 718x470; ColumnTextDate 'Дата'; ColumnTextAlarmState 'Статус'; ColumnTextAlarmText 'Аварийное сообщение'; ColumnTextTime 'Время'

screen "SIMATIC PLC system diagnostics" 800x480, template "Main"
   SysDiagControl "HmiScreenItemData" at 1,49 size 796x423
   Button "Back" at 1,1 size 159x47; TextOn 'Back'; TextOff 'Back'
      on Release: ActivateScreen("System screens", 0)

screen "System information" 800x480, template "Main"
   TextField "HmiScreenItemData" at 35,51 size 171x28; Text 'HMI device type:'
   TextField "HmiScreenItemData_1" at 241,51 size 524x28; Text 'KTP700 Basic+ PN 14.0.1.0'
   TextField "HmiScreenItemData_2" at 35,81 size 171x28; Text 'Connection:'
   TextField "HmiScreenItemData_3" at 241,81 size 524x28; Text 'PROFINET (X1)'
   TextField "HmiScreenItemData_4" at 35,111 size 171x28; Text 'PLC:'
   TextField "HmiScreenItemData_5" at 241,111 size 524x28; Text 'SIMATIC S7 1200'
   Button "Back" at 1,1 size 159x47; TextOn 'Back'; TextOff 'Back'
      on Release: ActivateScreen("System screens", 0)

screen "System screens" 800x480, template "Main"
   Button "Back" at 1,1 size 159x47; TextOn 'Back'; TextOff 'Back'
      on Release: ActivateScreen("Root screen", 0)
   Button "HmiScreenItemData" at 36,95 size 159x47; TextOn 'SIMATIC PLC system diagnos...'; TextOff 'SIMATIC PLC system diagnos...'; PictureOn "Navigates to SIMATIC PLC system diagnostics for KTP700 Basic+ PN 14.0.1.0"; PictureOff "Navigates to SIMATIC PLC system diagnostics for KTP700 Basic+ PN 14.0.1.0"
      on Release: ActivateScreen("SIMATIC PLC system diagnostics", 0)
   Button "HmiScreenItemData_1" at 36,154 size 159x47; TextOn 'Project information'; TextOff 'Project information'; PictureOn "Navigates to Project information for KTP700 Basic+ PN 14.0.1.0"; PictureOff "Navigates to Project information for KTP700 Basic+ PN 14.0.1.0"
      on Release: ActivateScreen("Project information", 0)
   Button "HmiScreenItemData_2" at 36,213 size 159x47; TextOn 'System information'; TextOff 'System information'; PictureOn "Navigates to System information for KTP700 Basic+ PN 14.0.1.0"; PictureOff "Navigates to System information for KTP700 Basic+ PN 14.0.1.0"
      on Release: ActivateScreen("System information", 0)
   Button "HmiScreenItemData_3" at 36,272 size 159x47; TextOn 'Different jobs'; TextOff 'Different jobs'; PictureOn "Navigates to Different jobs for KTP700 Basic+ PN 14.0.1.0"; PictureOff "Navigates to Different jobs for KTP700 Basic+ PN 14.0.1.0"
      on Release: ActivateScreen("Different jobs", 0)

screen "Different jobs" 800x480, template "Main"
   Button "Online" at 36,95 size 159x47; TextOn 'Online'; TextOff 'Online'
      on Release: function_bb44b551(0)
   Button "Offline" at 36,154 size 159x47; TextOn 'Offline'; TextOff 'Offline'
      on Release: function_bb44b551(1)
   Button "Transfer" at 36,213 size 159x47; TextOn 'Transfer'; TextOff 'Transfer'
      on Release: function_bb44b551(2)
   Button "Toggle language" at 36,272 size 159x47; TextOn 'Toggle language'; TextOff 'Toggle language'
      on Release: function_fb9197e8(-1)
   Button "Stop Runtime" at 36,331 size 159x47; TextOn 'Stop Runtime'; TextOff 'Stop Runtime'
      on Release: StopRuntime(0)
   Button "Back" at 1,1 size 159x47; TextOn 'Back'; TextOff 'Back'
      on Release: ActivateScreen("System screens", 0)

screen "Project information" 800x480, template "Main"
   TextField "HmiScreenItemData" at 35,51 size 171x28; Text 'Project name:'
   TextField "HmiScreenItemData_1" at 241,51 size 524x28; Text 'PolyMix_v0.1'
   TextField "HmiScreenItemData_2" at 35,81 size 171x28; Text 'Created on:'
   TextField "HmiScreenItemData_3" at 241,81 size 524x28; Text '10/24/2017 3:17:12 PM'
   TextField "HmiScreenItemData_4" at 35,111 size 171x28; Text 'Author:'
   TextField "HmiScreenItemData_5" at 241,111 size 524x28; Text 'WinCC'
   TextField "HmiScreenItemData_6" at 35,141 size 171x28; Text 'Description:'
   TextField "HmiScreenItemData_7" at 241,141 size 524x28; Text '(not configured)'
   Button "Back" at 1,1 size 159x47; TextOn 'Back'; TextOff 'Back'
      on Release: ActivateScreen("System screens", 0)

